(* Logix 5000 project; controller FV vendor 1 type 14 code 217 rev 31.11; software revision 31.00; part 18 of 63 *)
(* tags used below, declared in another part *)
   CheckTimeMask : INT;
   CWD : CHECKWORD_FLAGS;
   Delphi_Does_Eng_Func : BOOL;
   FR_AUDI1 : PlantItem;   // AUDI1
   FR_B240 : INT[255];   // DEBOUNCE Debounce Flags
   FR_BEACON1 : PlantItem;   // BEACON1
   FR_FV26_VA01 : PlantItem;   // FV26_VA01
   FR_FV27_VA01 : PlantItem;   // FV27_VA01
   FR_FV28_V : PlantItem;   // FV28_V
   FR_FV28_VA01 : PlantItem;   // FV28_VA01
   FR_FVS_P01 : PlantItem;   // FVS_P01
   FR_N14 : INT[265];   // MVFV CIP Comms to MVFV CIP Un it PLC
   FR_N140 : INT[265];   // CIP
   FR_N255 : INT[265];   // CHECKWORDS
   FR_N26 : INT[265];   // FV26
   FR_N27 : INT[265];   // FV27
   FR_N28 : INT[265];   // FV28
   FR_N29 : INT[265];   // FV29
   FR_N30 : INT[265];   // FV30
   FR_N31 : INT[265];   // FV31
   FR_N99 : INT[265];   // COMMENT Comment Lines
   FR_R3_SW3_1 : PlantItem;   // R3_SW3_1
   FR_R3_SW3_2 : PlantItem;   // R3_SW3_2
   FR_R3_SW3_3 : PlantItem;   // R3_SW3_3
   FR_T144 : TIMER[255];   // CIP
   FR_VB4_AV20 : PlantItem;   // VB4_AV20
   FR_VB4_AV22 : PlantItem;   // VB4_AV22
   FR_YP1_CIP : PlantItem;   // YP1_CIP
   FR_YP2_CIP : PlantItem;   // YP2_CIP
   FR_YP3_CIP : PlantItem;   // YP3_CIP
   TempChecktime : DINT;
(* FR_Common, continued *)

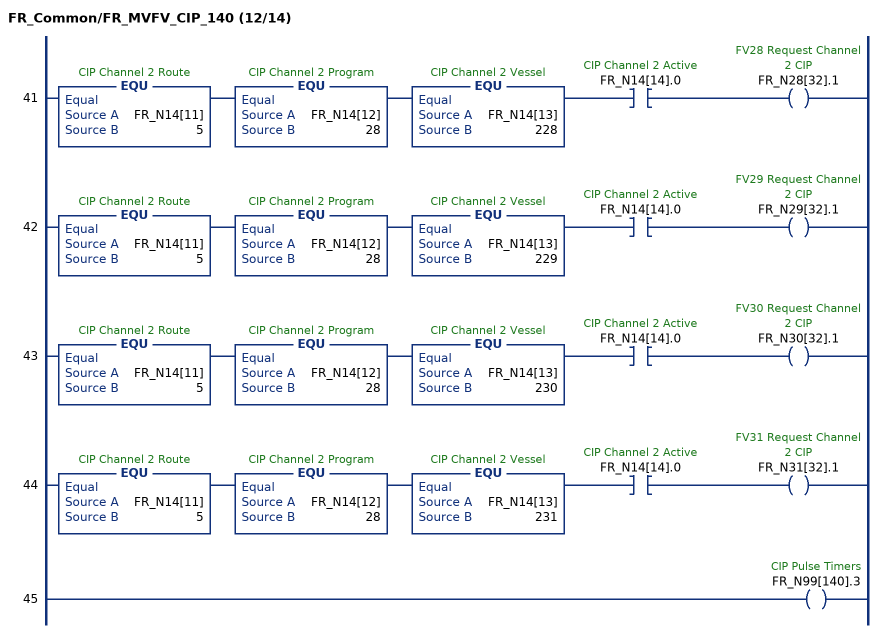
   [picture p297: FR_Common/FR_MVFV_CIP_140 rungs 41-45]
   41: EQU(FR_N14[11],5)EQU(FR_N14[12],28)EQU(FR_N14[13],228)XIC(FR_N14[14].0)OTE(FR_N28[32].1);
   42: EQU(FR_N14[11],5)EQU(FR_N14[12],28)EQU(FR_N14[13],229)XIC(FR_N14[14].0)OTE(FR_N29[32].1);
   43: EQU(FR_N14[11],5)EQU(FR_N14[12],28)EQU(FR_N14[13],230)XIC(FR_N14[14].0)OTE(FR_N30[32].1);
   44: EQU(FR_N14[11],5)EQU(FR_N14[12],28)EQU(FR_N14[13],231)XIC(FR_N14[14].0)OTE(FR_N31[32].1);
   45: OTE(FR_N99[140].3);
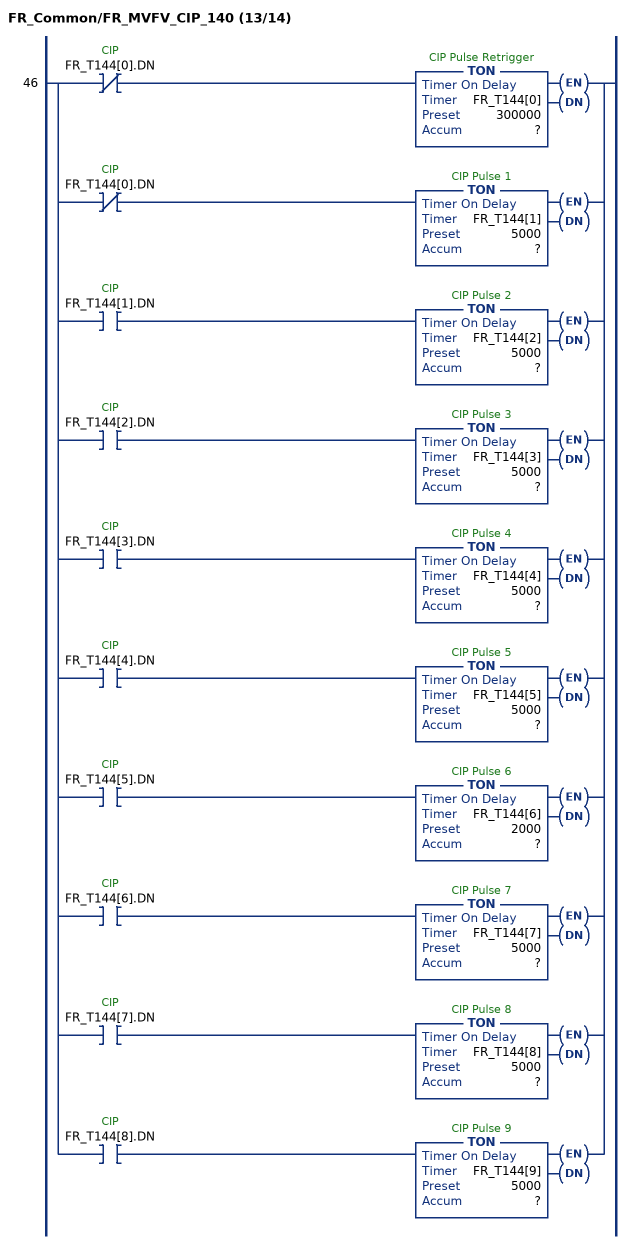
   46: [XIO(FR_T144[0].DN) TON(FR_T144[0],?,?) ,XIO(FR_T144[0].DN) TON(FR_T144[1],?,?) ,XIC(FR_T144[1].DN) TON(FR_T144[2],?,?) ,XIC(FR_T144[2].DN) TON(FR_T144[3],?,?) ,XIC(FR_T144[3].DN) TON(FR_T144[4],?,?) ,XIC(FR_T144[4].DN) TON(FR_T144[5],?,?) ,XIC(FR_T144[5].DN) TON(FR_T144[6],?,?) ,XIC(FR_T144[6].DN) TON(FR_T144[7],?,?) ,XIC(FR_T144[7].DN) TON(FR_T144[8],?,?) ,XIC(FR_T144[8].DN) TON(FR_T144[9],?,?) ];
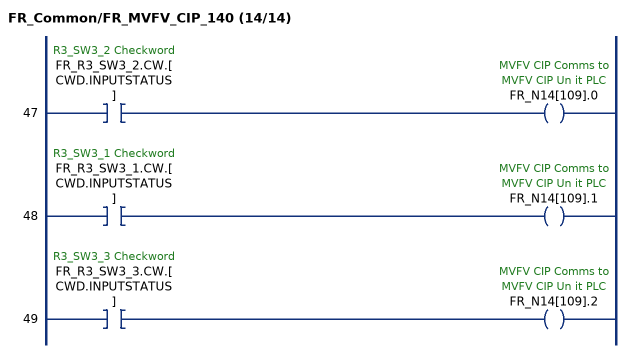
   47: XIC(FR_R3_SW3_2.CW.[CWD.INPUTSTATUS])OTE(FR_N14[109].0);
   48: XIC(FR_R3_SW3_1.CW.[CWD.INPUTSTATUS])OTE(FR_N14[109].1);
   49: XIC(FR_R3_SW3_3.CW.[CWD.INPUTSTATUS])OTE(FR_N14[109].2);
END_ROUTINE

ROUTINE FR_MVFV_CIP_O_141   (* ladder *)
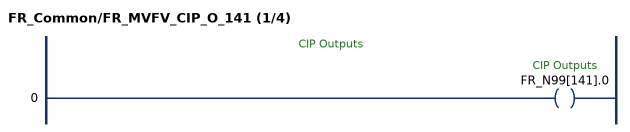
   // CIP Outputs
   0: OTE(FR_N99[141].0);
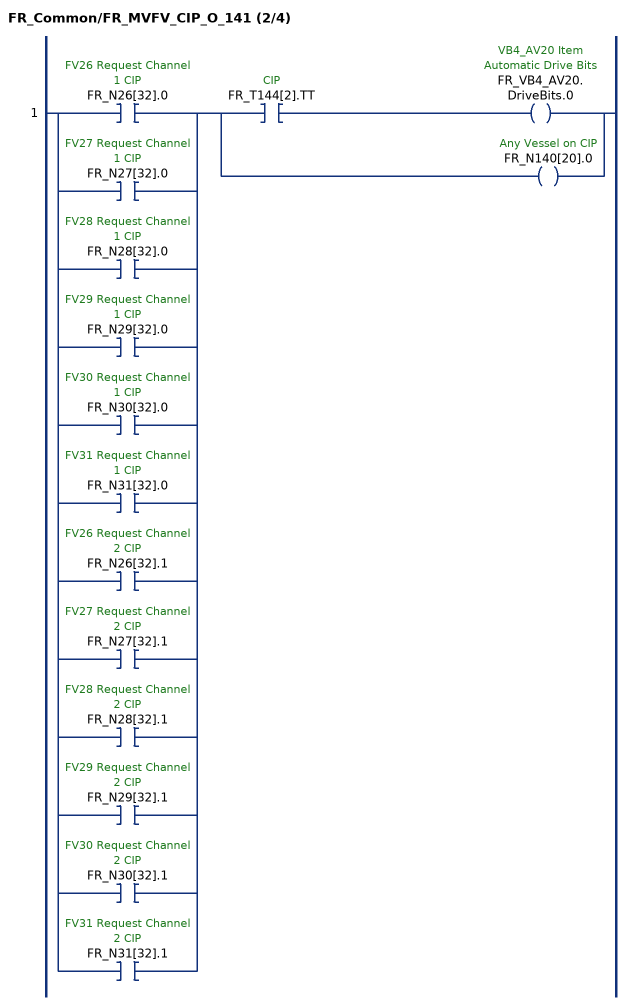
   1: [XIC(FR_N26[32].0) ,XIC(FR_N27[32].0) ,XIC(FR_N28[32].0) ,XIC(FR_N29[32].0) ,XIC(FR_N30[32].0) ,XIC(FR_N31[32].0) ,XIC(FR_N26[32].1) ,XIC(FR_N27[32].1) ,XIC(FR_N28[32].1) ,XIC(FR_N29[32].1) ,XIC(FR_N30[32].1) ,XIC(FR_N31[32].1) ][XIC(FR_T144[2].TT) OTE(FR_VB4_AV20.DriveBits.0) ,OTE(FR_N140[20].0) ];
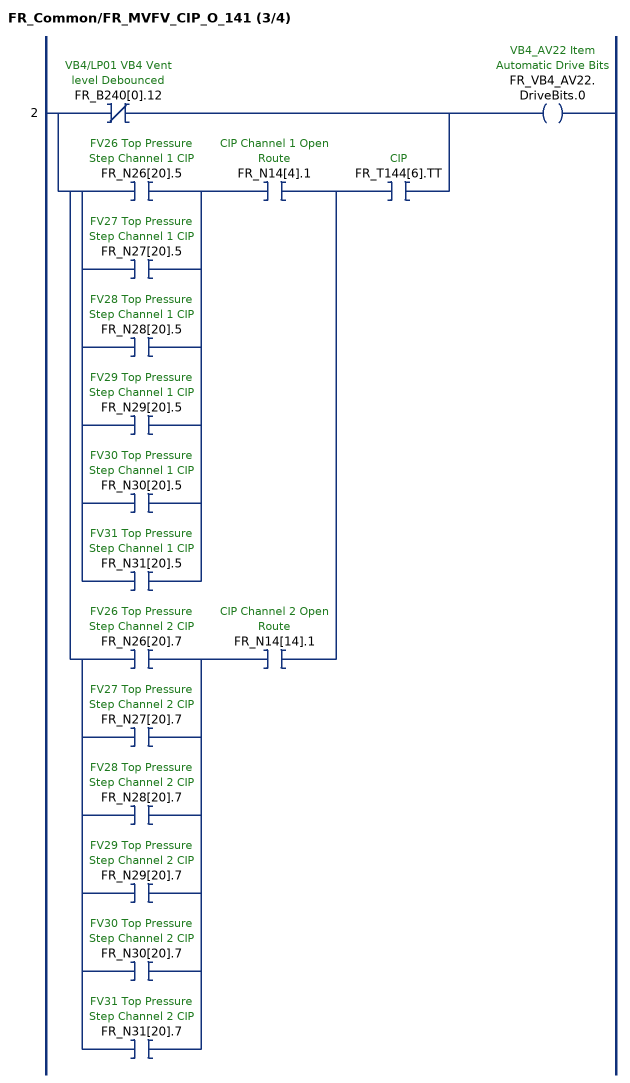
   2: [XIO(FR_B240[0].12) ,[[XIC(FR_N26[20].5) ,XIC(FR_N27[20].5) ,XIC(FR_N28[20].5) ,XIC(FR_N29[20].5) ,XIC(FR_N30[20].5) ,XIC(FR_N31[20].5) ] XIC(FR_N14[4].1) ,[XIC(FR_N26[20].7) ,XIC(FR_N27[20].7) ,XIC(FR_N28[20].7) ,XIC(FR_N29[20].7) ,XIC(FR_N30[20].7) ,XIC(FR_N31[20].7) ] XIC(FR_N14[14].1) ] XIC(FR_T144[6].TT) ]OTE(FR_VB4_AV22.DriveBits.0);
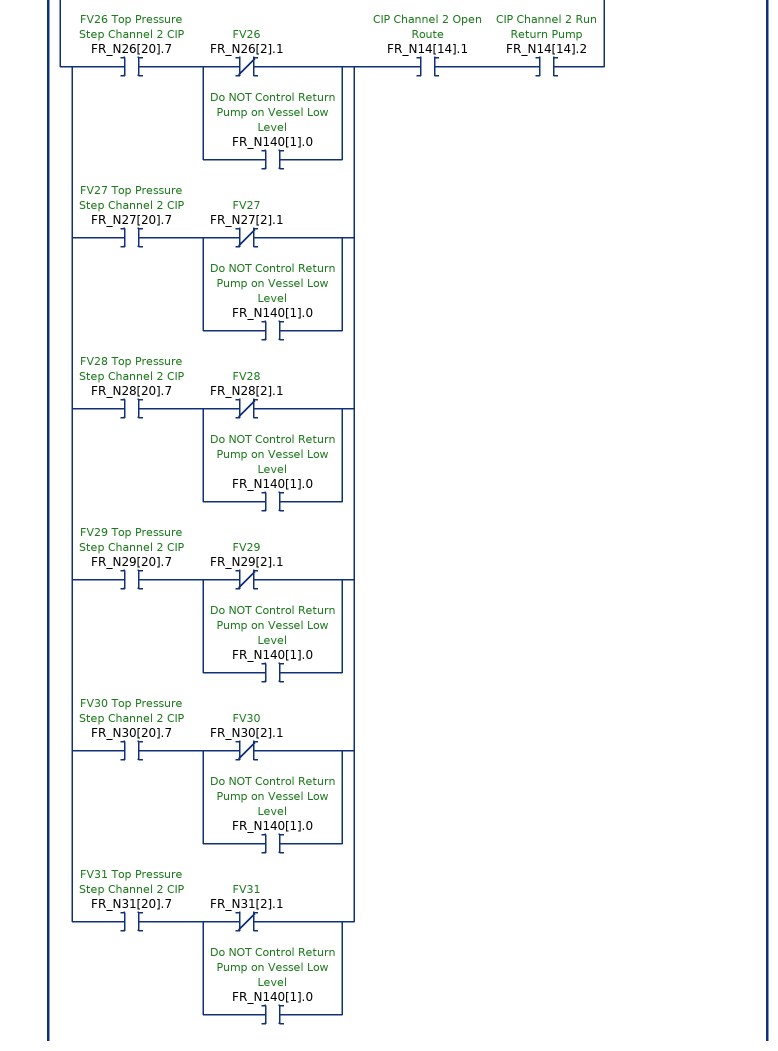
   3: [[XIC(FR_N26[20].5) [XIO(FR_N26[2].1) ,XIC(FR_N140[1].0) ] ,XIC(FR_N27[20].5) [XIO(FR_N27[2].1) ,XIC(FR_N140[1].0) ] ,XIC(FR_N28[20].5) [XIO(FR_N28[2].1) ,XIC(FR_N140[1].0) ] ,XIC(FR_N29[20].5) [XIO(FR_N29[2].1) ,XIC(FR_N140[1].0) ] ,XIC(FR_N30[20].5) [XIO(FR_N30[2].1) ,XIC(FR_N140[1].0) ] ,XIC(FR_N31[20].5) [XIO(FR_N31[2].1) ,XIC(FR_N140[1].0) ] ] XIC(FR_N14[4].1) XIC(FR_N14[4].2) ,[XIC(FR_N26[20].7) [XIO(FR_N26[2].1) ,XIC(FR_N140[1].0) ] ,XIC(FR_N27[20].7) [XIO(FR_N27[2].1) ,XIC(FR_N140[1].0) ] ,XIC(FR_N28[20].7) [XIO(FR_N28[2].1) ,XIC(FR_N140[1].0) ] ,XIC(FR_N29[20].7) [XIO(FR_N29[2].1) ,XIC(FR_N140[1].0) ] ,XIC(FR_N30[20].7) [XIO(FR_N30[2].1) ,XIC(FR_N140[1].0) ] ,XIC(FR_N31[20].7) [XIO(FR_N31[2].1) ,XIC(FR_N140[1].0) ] ] XIC(FR_N14[14].1) XIC(FR_N14[14].2) ]OTE(FR_FVS_P01.DriveBits.0);
END_ROUTINE

ROUTINE FR_Old_Checkword_Relaying   (* ladder *)
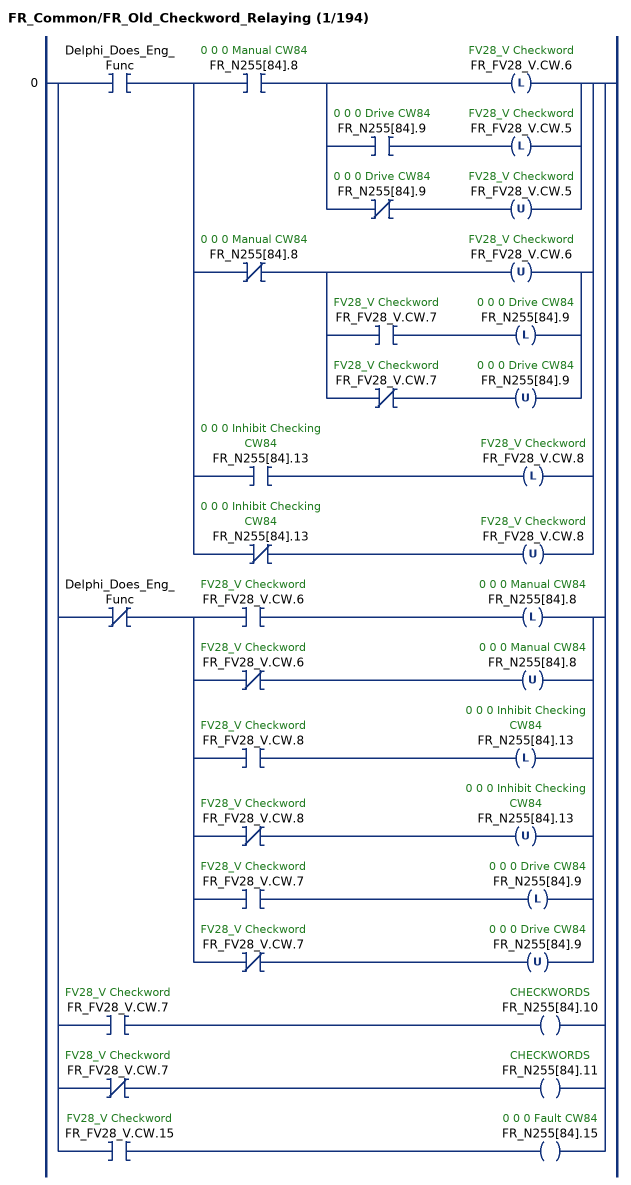
   0: [XIC(Delphi_Does_Eng_Func) [[XIC(FR_N255[84].8) [OTL(FR_FV28_V.CW.6) ,XIC(FR_N255[84].9) OTL(FR_FV28_V.CW.5) ,XIO(FR_N255[84].9) OTU(FR_FV28_V.CW.5) ] ,XIO(FR_N255[84].8) [OTU(FR_FV28_V.CW.6) ,[XIC(FR_FV28_V.CW.7) OTL(FR_N255[84].9) ,XIO(FR_FV28_V.CW.7) OTU(FR_N255[84].9) ] ] ] ,[XIC(FR_N255[84].13) OTL(FR_FV28_V.CW.8) ,XIO(FR_N255[84].13) OTU(FR_FV28_V.CW.8) ] ] ,XIO(Delphi_Does_Eng_Func) [[XIC(FR_FV28_V.CW.6) OTL(FR_N255[84].8) ,XIO(FR_FV28_V.CW.6) OTU(FR_N255[84].8) ] ,[XIC(FR_FV28_V.CW.8) OTL(FR_N255[84].13) ,XIO(FR_FV28_V.CW.8) OTU(FR_N255[84].13) ] ,[XIC(FR_FV28_V.CW.7) OTL(FR_N255[84].9) ,XIO(FR_FV28_V.CW.7) OTU(FR_N255[84].9) ] ] ,XIC(FR_FV28_V.CW.7) OTE(FR_N255[84].10) ,XIO(FR_FV28_V.CW.7) OTE(FR_N255[84].11) ,XIC(FR_FV28_V.CW.15) OTE(FR_N255[84].15) ];
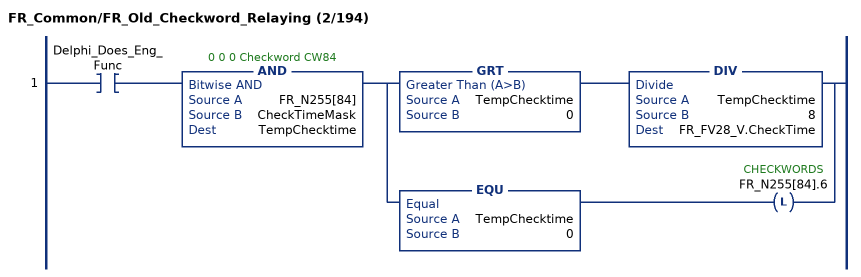
   1: XIC(Delphi_Does_Eng_Func)AND(FR_N255[84],CheckTimeMask,TempChecktime)[GRT(TempChecktime,0) DIV(TempChecktime,8,FR_FV28_V.CheckTime) ,EQU(TempChecktime,0) OTL(FR_N255[84].6) ];
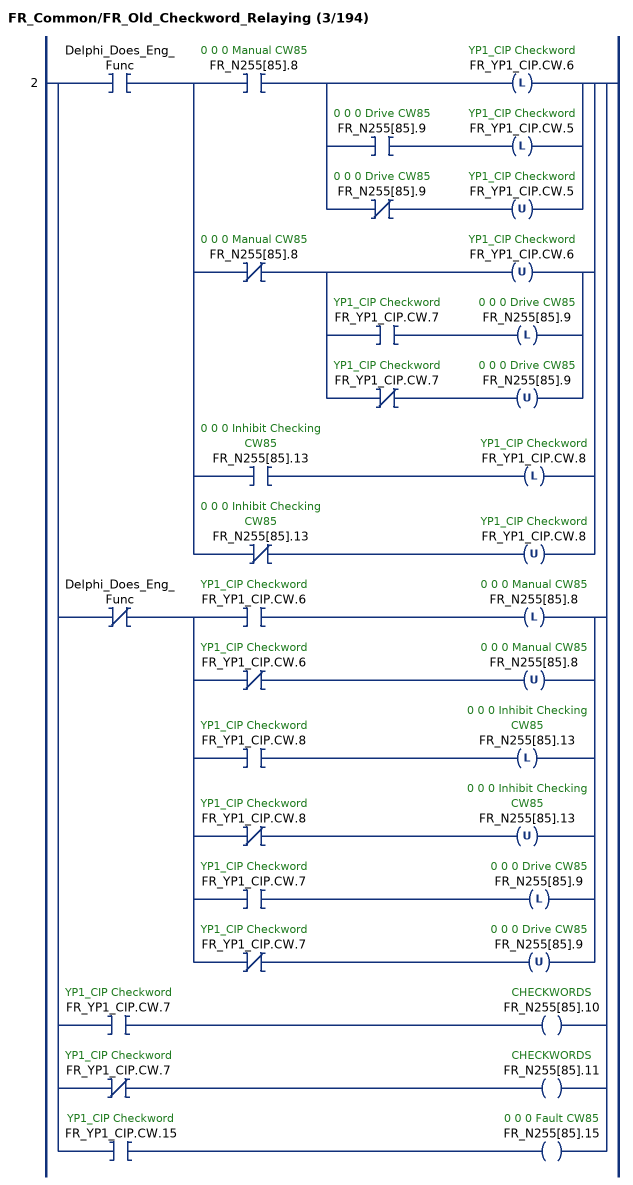
   2: [XIC(Delphi_Does_Eng_Func) [[XIC(FR_N255[85].8) [OTL(FR_YP1_CIP.CW.6) ,XIC(FR_N255[85].9) OTL(FR_YP1_CIP.CW.5) ,XIO(FR_N255[85].9) OTU(FR_YP1_CIP.CW.5) ] ,XIO(FR_N255[85].8) [OTU(FR_YP1_CIP.CW.6) ,[XIC(FR_YP1_CIP.CW.7) OTL(FR_N255[85].9) ,XIO(FR_YP1_CIP.CW.7) OTU(FR_N255[85].9) ] ] ] ,[XIC(FR_N255[85].13) OTL(FR_YP1_CIP.CW.8) ,XIO(FR_N255[85].13) OTU(FR_YP1_CIP.CW.8) ] ] ,XIO(Delphi_Does_Eng_Func) [[XIC(FR_YP1_CIP.CW.6) OTL(FR_N255[85].8) ,XIO(FR_YP1_CIP.CW.6) OTU(FR_N255[85].8) ] ,[XIC(FR_YP1_CIP.CW.8) OTL(FR_N255[85].13) ,XIO(FR_YP1_CIP.CW.8) OTU(FR_N255[85].13) ] ,[XIC(FR_YP1_CIP.CW.7) OTL(FR_N255[85].9) ,XIO(FR_YP1_CIP.CW.7) OTU(FR_N255[85].9) ] ] ,XIC(FR_YP1_CIP.CW.7) OTE(FR_N255[85].10) ,XIO(FR_YP1_CIP.CW.7) OTE(FR_N255[85].11) ,XIC(FR_YP1_CIP.CW.15) OTE(FR_N255[85].15) ];
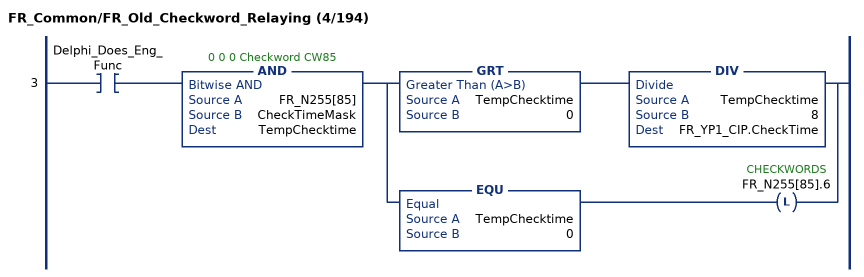
   3: XIC(Delphi_Does_Eng_Func)AND(FR_N255[85],CheckTimeMask,TempChecktime)[GRT(TempChecktime,0) DIV(TempChecktime,8,FR_YP1_CIP.CheckTime) ,EQU(TempChecktime,0) OTL(FR_N255[85].6) ];
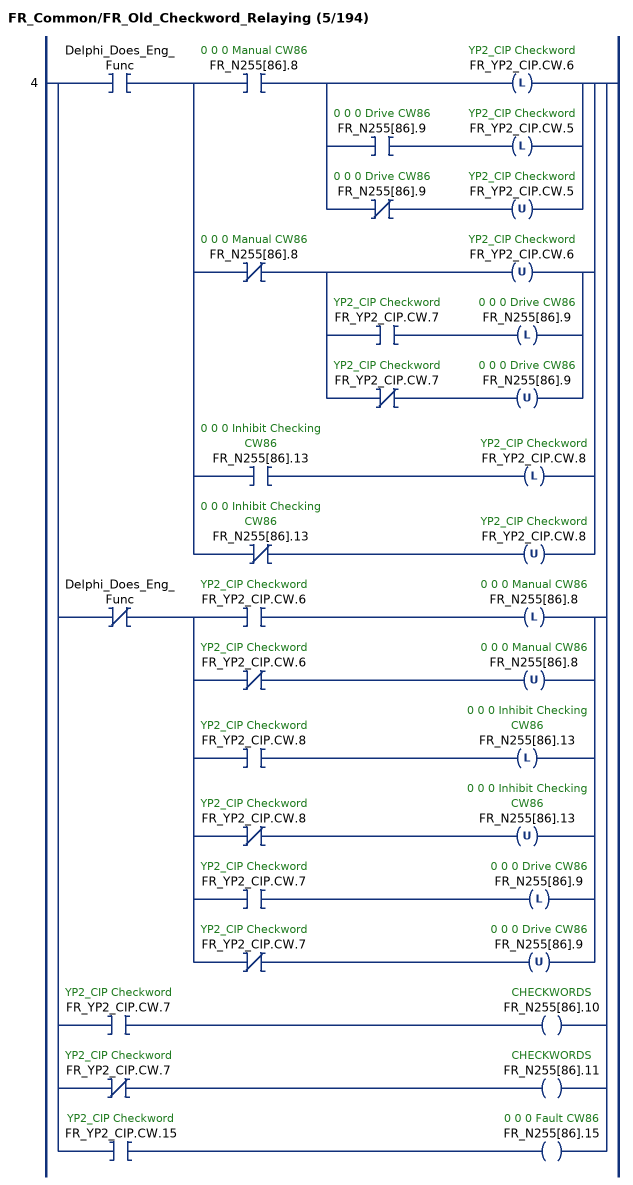
   4: [XIC(Delphi_Does_Eng_Func) [[XIC(FR_N255[86].8) [OTL(FR_YP2_CIP.CW.6) ,XIC(FR_N255[86].9) OTL(FR_YP2_CIP.CW.5) ,XIO(FR_N255[86].9) OTU(FR_YP2_CIP.CW.5) ] ,XIO(FR_N255[86].8) [OTU(FR_YP2_CIP.CW.6) ,[XIC(FR_YP2_CIP.CW.7) OTL(FR_N255[86].9) ,XIO(FR_YP2_CIP.CW.7) OTU(FR_N255[86].9) ] ] ] ,[XIC(FR_N255[86].13) OTL(FR_YP2_CIP.CW.8) ,XIO(FR_N255[86].13) OTU(FR_YP2_CIP.CW.8) ] ] ,XIO(Delphi_Does_Eng_Func) [[XIC(FR_YP2_CIP.CW.6) OTL(FR_N255[86].8) ,XIO(FR_YP2_CIP.CW.6) OTU(FR_N255[86].8) ] ,[XIC(FR_YP2_CIP.CW.8) OTL(FR_N255[86].13) ,XIO(FR_YP2_CIP.CW.8) OTU(FR_N255[86].13) ] ,[XIC(FR_YP2_CIP.CW.7) OTL(FR_N255[86].9) ,XIO(FR_YP2_CIP.CW.7) OTU(FR_N255[86].9) ] ] ,XIC(FR_YP2_CIP.CW.7) OTE(FR_N255[86].10) ,XIO(FR_YP2_CIP.CW.7) OTE(FR_N255[86].11) ,XIC(FR_YP2_CIP.CW.15) OTE(FR_N255[86].15) ];
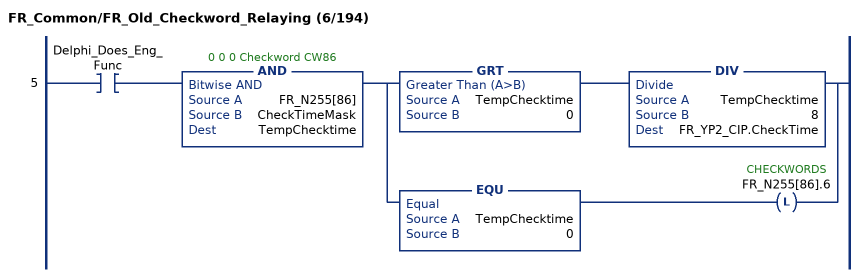
   5: XIC(Delphi_Does_Eng_Func)AND(FR_N255[86],CheckTimeMask,TempChecktime)[GRT(TempChecktime,0) DIV(TempChecktime,8,FR_YP2_CIP.CheckTime) ,EQU(TempChecktime,0) OTL(FR_N255[86].6) ];
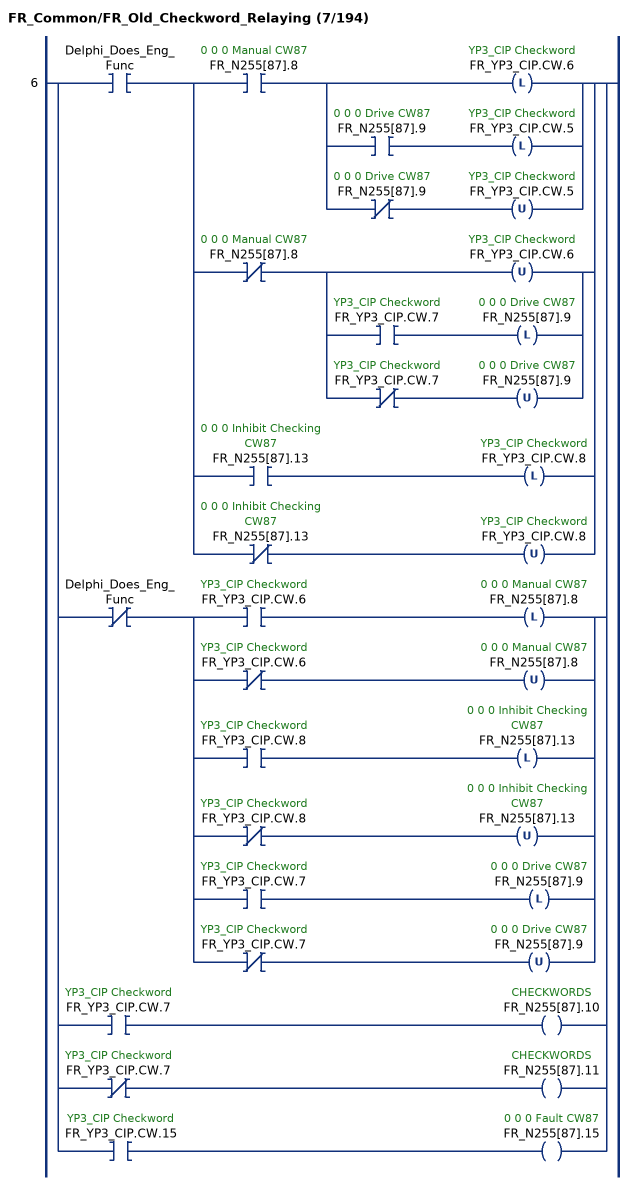
   6: [XIC(Delphi_Does_Eng_Func) [[XIC(FR_N255[87].8) [OTL(FR_YP3_CIP.CW.6) ,XIC(FR_N255[87].9) OTL(FR_YP3_CIP.CW.5) ,XIO(FR_N255[87].9) OTU(FR_YP3_CIP.CW.5) ] ,XIO(FR_N255[87].8) [OTU(FR_YP3_CIP.CW.6) ,[XIC(FR_YP3_CIP.CW.7) OTL(FR_N255[87].9) ,XIO(FR_YP3_CIP.CW.7) OTU(FR_N255[87].9) ] ] ] ,[XIC(FR_N255[87].13) OTL(FR_YP3_CIP.CW.8) ,XIO(FR_N255[87].13) OTU(FR_YP3_CIP.CW.8) ] ] ,XIO(Delphi_Does_Eng_Func) [[XIC(FR_YP3_CIP.CW.6) OTL(FR_N255[87].8) ,XIO(FR_YP3_CIP.CW.6) OTU(FR_N255[87].8) ] ,[XIC(FR_YP3_CIP.CW.8) OTL(FR_N255[87].13) ,XIO(FR_YP3_CIP.CW.8) OTU(FR_N255[87].13) ] ,[XIC(FR_YP3_CIP.CW.7) OTL(FR_N255[87].9) ,XIO(FR_YP3_CIP.CW.7) OTU(FR_N255[87].9) ] ] ,XIC(FR_YP3_CIP.CW.7) OTE(FR_N255[87].10) ,XIO(FR_YP3_CIP.CW.7) OTE(FR_N255[87].11) ,XIC(FR_YP3_CIP.CW.15) OTE(FR_N255[87].15) ];
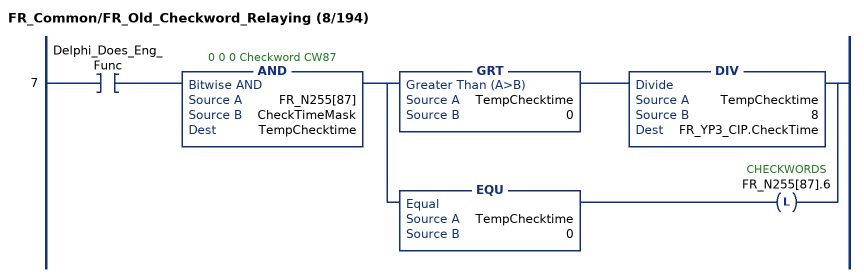
   7: XIC(Delphi_Does_Eng_Func)AND(FR_N255[87],CheckTimeMask,TempChecktime)[GRT(TempChecktime,0) DIV(TempChecktime,8,FR_YP3_CIP.CheckTime) ,EQU(TempChecktime,0) OTL(FR_N255[87].6) ];
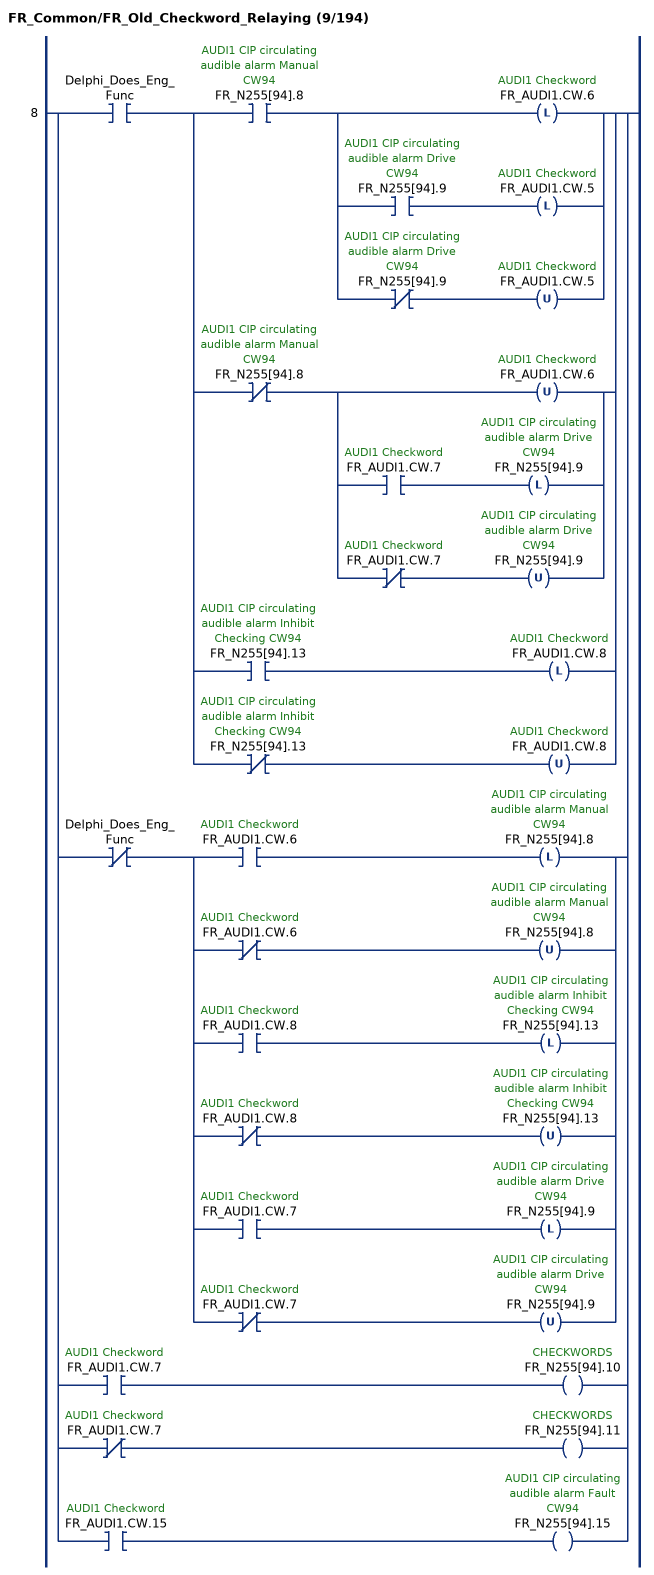
   8: [XIC(Delphi_Does_Eng_Func) [[XIC(FR_N255[94].8) [OTL(FR_AUDI1.CW.6) ,XIC(FR_N255[94].9) OTL(FR_AUDI1.CW.5) ,XIO(FR_N255[94].9) OTU(FR_AUDI1.CW.5) ] ,XIO(FR_N255[94].8) [OTU(FR_AUDI1.CW.6) ,[XIC(FR_AUDI1.CW.7) OTL(FR_N255[94].9) ,XIO(FR_AUDI1.CW.7) OTU(FR_N255[94].9) ] ] ] ,[XIC(FR_N255[94].13) OTL(FR_AUDI1.CW.8) ,XIO(FR_N255[94].13) OTU(FR_AUDI1.CW.8) ] ] ,XIO(Delphi_Does_Eng_Func) [[XIC(FR_AUDI1.CW.6) OTL(FR_N255[94].8) ,XIO(FR_AUDI1.CW.6) OTU(FR_N255[94].8) ] ,[XIC(FR_AUDI1.CW.8) OTL(FR_N255[94].13) ,XIO(FR_AUDI1.CW.8) OTU(FR_N255[94].13) ] ,[XIC(FR_AUDI1.CW.7) OTL(FR_N255[94].9) ,XIO(FR_AUDI1.CW.7) OTU(FR_N255[94].9) ] ] ,XIC(FR_AUDI1.CW.7) OTE(FR_N255[94].10) ,XIO(FR_AUDI1.CW.7) OTE(FR_N255[94].11) ,XIC(FR_AUDI1.CW.15) OTE(FR_N255[94].15) ];
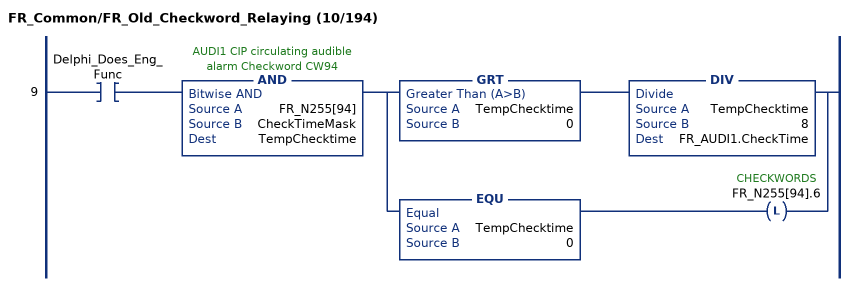
   9: XIC(Delphi_Does_Eng_Func)AND(FR_N255[94],CheckTimeMask,TempChecktime)[GRT(TempChecktime,0) DIV(TempChecktime,8,FR_AUDI1.CheckTime) ,EQU(TempChecktime,0) OTL(FR_N255[94].6) ];
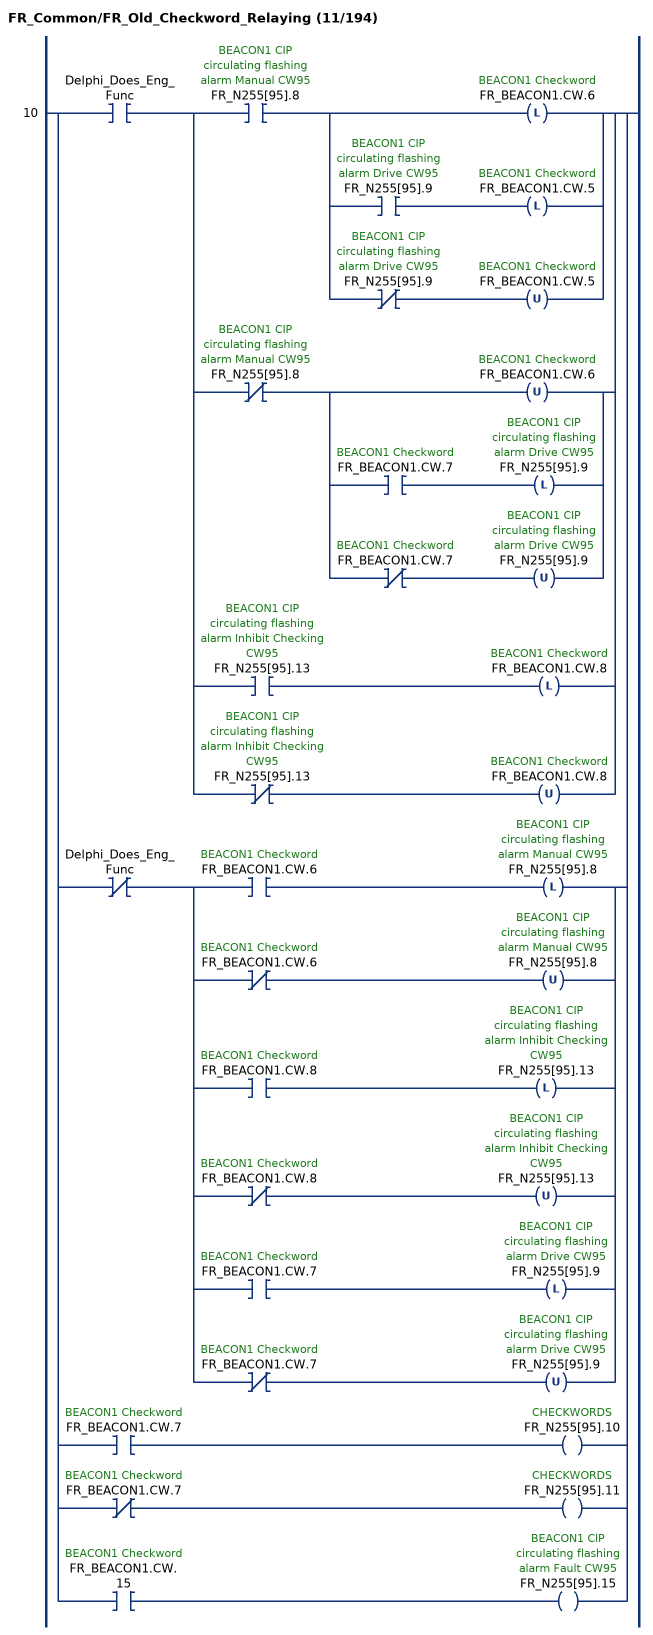
   10: [XIC(Delphi_Does_Eng_Func) [[XIC(FR_N255[95].8) [OTL(FR_BEACON1.CW.6) ,XIC(FR_N255[95].9) OTL(FR_BEACON1.CW.5) ,XIO(FR_N255[95].9) OTU(FR_BEACON1.CW.5) ] ,XIO(FR_N255[95].8) [OTU(FR_BEACON1.CW.6) ,[XIC(FR_BEACON1.CW.7) OTL(FR_N255[95].9) ,XIO(FR_BEACON1.CW.7) OTU(FR_N255[95].9) ] ] ] ,[XIC(FR_N255[95].13) OTL(FR_BEACON1.CW.8) ,XIO(FR_N255[95].13) OTU(FR_BEACON1.CW.8) ] ] ,XIO(Delphi_Does_Eng_Func) [[XIC(FR_BEACON1.CW.6) OTL(FR_N255[95].8) ,XIO(FR_BEACON1.CW.6) OTU(FR_N255[95].8) ] ,[XIC(FR_BEACON1.CW.8) OTL(FR_N255[95].13) ,XIO(FR_BEACON1.CW.8) OTU(FR_N255[95].13) ] ,[XIC(FR_BEACON1.CW.7) OTL(FR_N255[95].9) ,XIO(FR_BEACON1.CW.7) OTU(FR_N255[95].9) ] ] ,XIC(FR_BEACON1.CW.7) OTE(FR_N255[95].10) ,XIO(FR_BEACON1.CW.7) OTE(FR_N255[95].11) ,XIC(FR_BEACON1.CW.15) OTE(FR_N255[95].15) ];
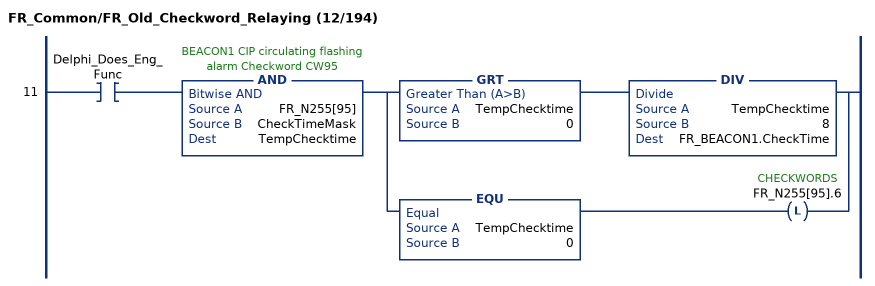
   11: XIC(Delphi_Does_Eng_Func)AND(FR_N255[95],CheckTimeMask,TempChecktime)[GRT(TempChecktime,0) DIV(TempChecktime,8,FR_BEACON1.CheckTime) ,EQU(TempChecktime,0) OTL(FR_N255[95].6) ];
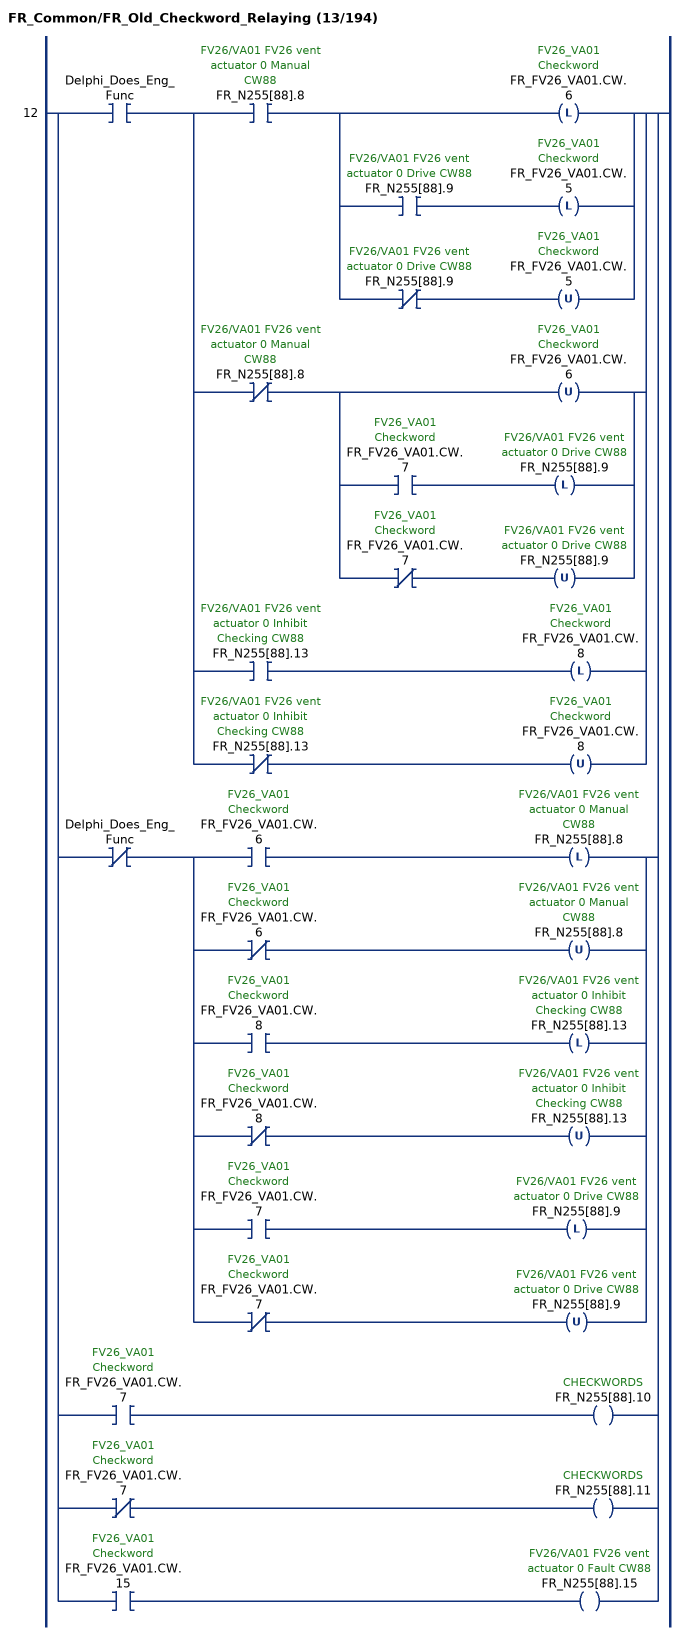
   12: [XIC(Delphi_Does_Eng_Func) [[XIC(FR_N255[88].8) [OTL(FR_FV26_VA01.CW.6) ,XIC(FR_N255[88].9) OTL(FR_FV26_VA01.CW.5) ,XIO(FR_N255[88].9) OTU(FR_FV26_VA01.CW.5) ] ,XIO(FR_N255[88].8) [OTU(FR_FV26_VA01.CW.6) ,[XIC(FR_FV26_VA01.CW.7) OTL(FR_N255[88].9) ,XIO(FR_FV26_VA01.CW.7) OTU(FR_N255[88].9) ] ] ] ,[XIC(FR_N255[88].13) OTL(FR_FV26_VA01.CW.8) ,XIO(FR_N255[88].13) OTU(FR_FV26_VA01.CW.8) ] ] ,XIO(Delphi_Does_Eng_Func) [[XIC(FR_FV26_VA01.CW.6) OTL(FR_N255[88].8) ,XIO(FR_FV26_VA01.CW.6) OTU(FR_N255[88].8) ] ,[XIC(FR_FV26_VA01.CW.8) OTL(FR_N255[88].13) ,XIO(FR_FV26_VA01.CW.8) OTU(FR_N255[88].13) ] ,[XIC(FR_FV26_VA01.CW.7) OTL(FR_N255[88].9) ,XIO(FR_FV26_VA01.CW.7) OTU(FR_N255[88].9) ] ] ,XIC(FR_FV26_VA01.CW.7) OTE(FR_N255[88].10) ,XIO(FR_FV26_VA01.CW.7) OTE(FR_N255[88].11) ,XIC(FR_FV26_VA01.CW.15) OTE(FR_N255[88].15) ];
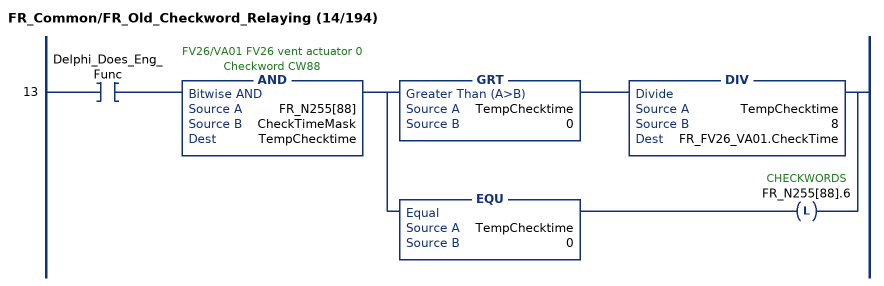
   13: XIC(Delphi_Does_Eng_Func)AND(FR_N255[88],CheckTimeMask,TempChecktime)[GRT(TempChecktime,0) DIV(TempChecktime,8,FR_FV26_VA01.CheckTime) ,EQU(TempChecktime,0) OTL(FR_N255[88].6) ];
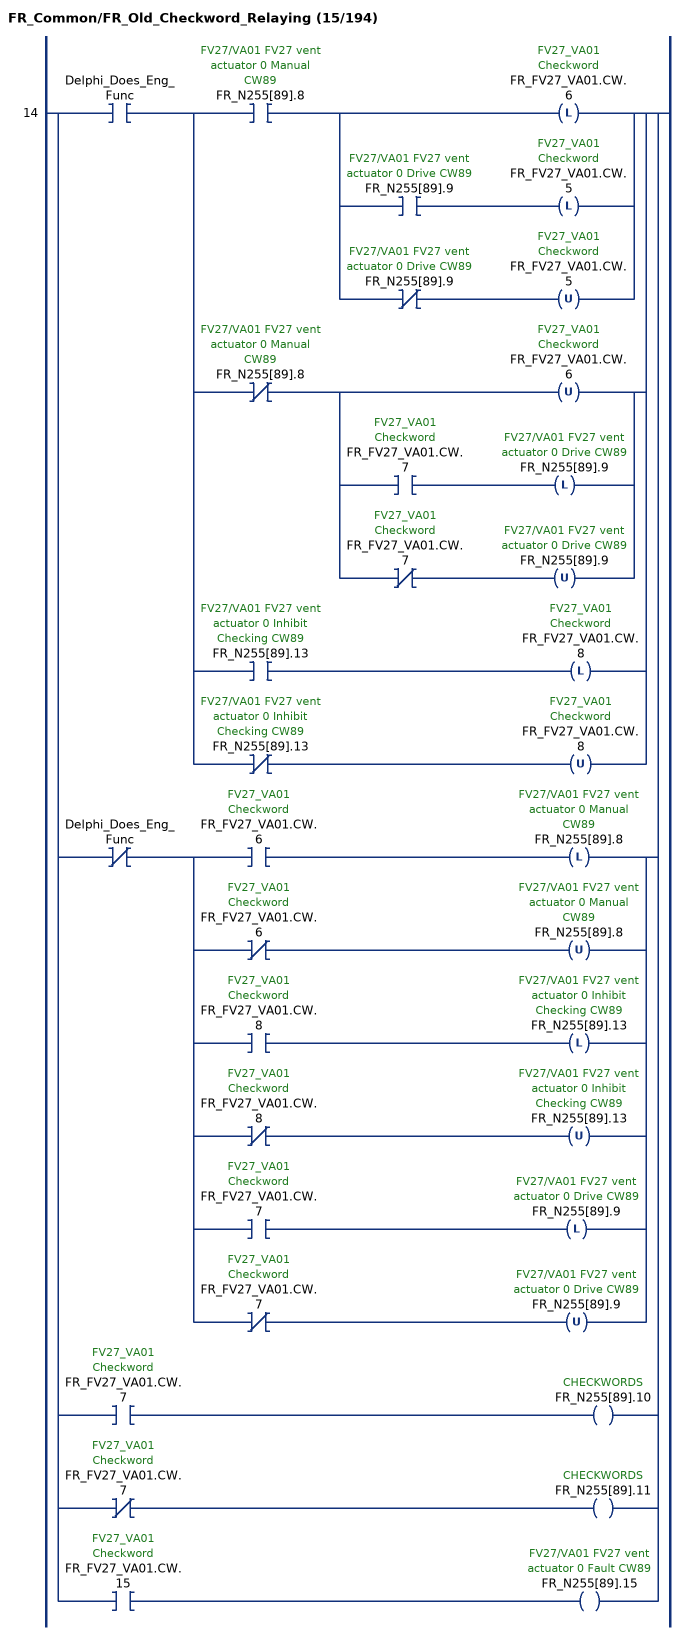
   14: [XIC(Delphi_Does_Eng_Func) [[XIC(FR_N255[89].8) [OTL(FR_FV27_VA01.CW.6) ,XIC(FR_N255[89].9) OTL(FR_FV27_VA01.CW.5) ,XIO(FR_N255[89].9) OTU(FR_FV27_VA01.CW.5) ] ,XIO(FR_N255[89].8) [OTU(FR_FV27_VA01.CW.6) ,[XIC(FR_FV27_VA01.CW.7) OTL(FR_N255[89].9) ,XIO(FR_FV27_VA01.CW.7) OTU(FR_N255[89].9) ] ] ] ,[XIC(FR_N255[89].13) OTL(FR_FV27_VA01.CW.8) ,XIO(FR_N255[89].13) OTU(FR_FV27_VA01.CW.8) ] ] ,XIO(Delphi_Does_Eng_Func) [[XIC(FR_FV27_VA01.CW.6) OTL(FR_N255[89].8) ,XIO(FR_FV27_VA01.CW.6) OTU(FR_N255[89].8) ] ,[XIC(FR_FV27_VA01.CW.8) OTL(FR_N255[89].13) ,XIO(FR_FV27_VA01.CW.8) OTU(FR_N255[89].13) ] ,[XIC(FR_FV27_VA01.CW.7) OTL(FR_N255[89].9) ,XIO(FR_FV27_VA01.CW.7) OTU(FR_N255[89].9) ] ] ,XIC(FR_FV27_VA01.CW.7) OTE(FR_N255[89].10) ,XIO(FR_FV27_VA01.CW.7) OTE(FR_N255[89].11) ,XIC(FR_FV27_VA01.CW.15) OTE(FR_N255[89].15) ];
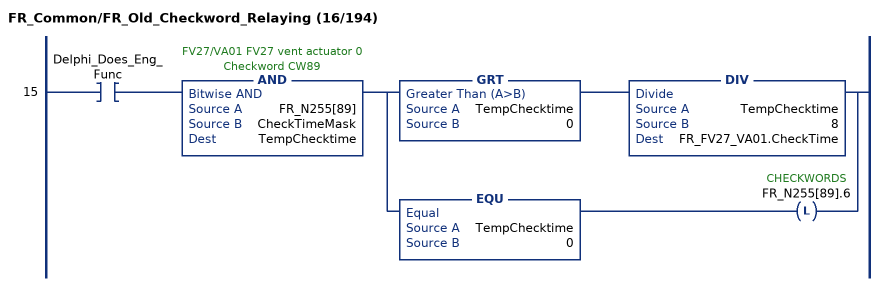
   15: XIC(Delphi_Does_Eng_Func)AND(FR_N255[89],CheckTimeMask,TempChecktime)[GRT(TempChecktime,0) DIV(TempChecktime,8,FR_FV27_VA01.CheckTime) ,EQU(TempChecktime,0) OTL(FR_N255[89].6) ];
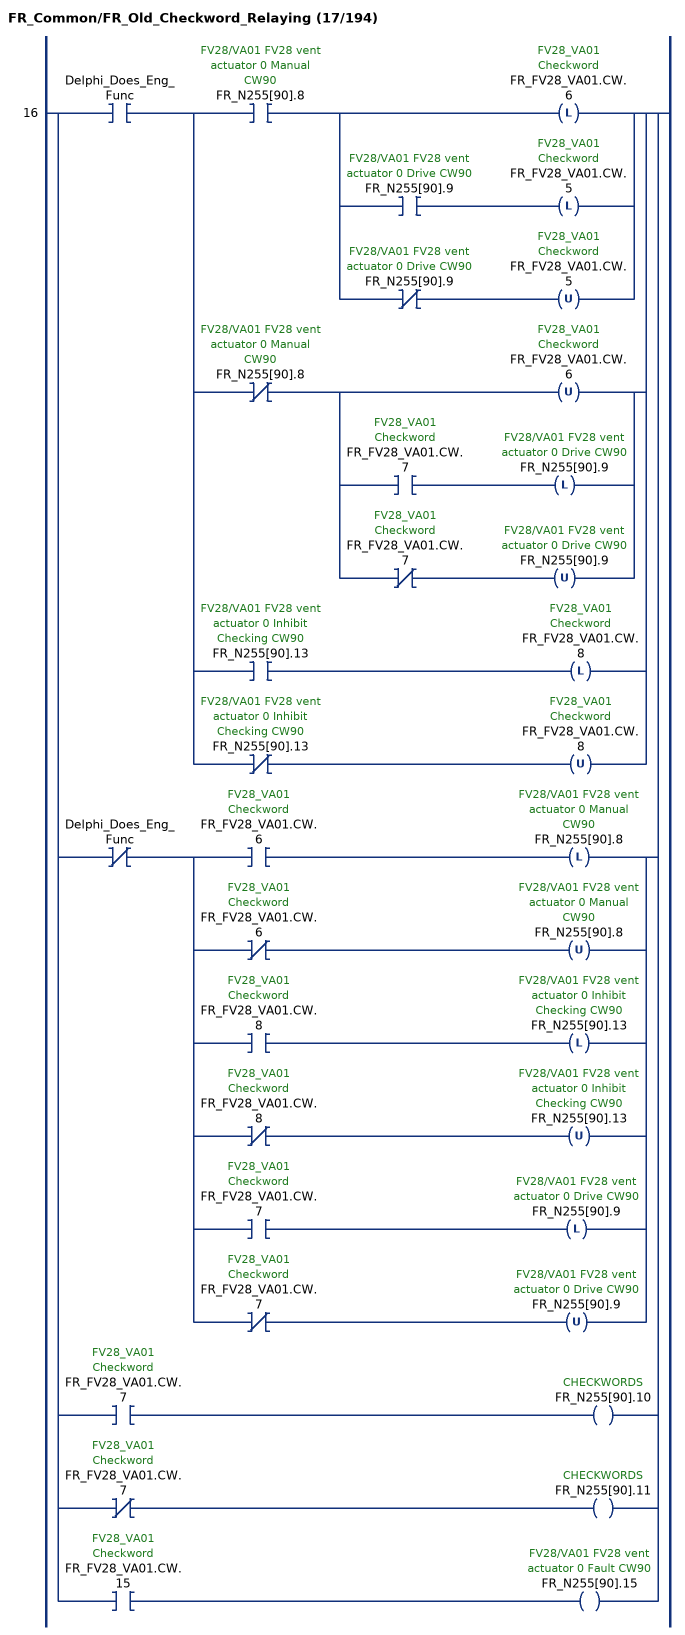
   16: [XIC(Delphi_Does_Eng_Func) [[XIC(FR_N255[90].8) [OTL(FR_FV28_VA01.CW.6) ,XIC(FR_N255[90].9) OTL(FR_FV28_VA01.CW.5) ,XIO(FR_N255[90].9) OTU(FR_FV28_VA01.CW.5) ] ,XIO(FR_N255[90].8) [OTU(FR_FV28_VA01.CW.6) ,[XIC(FR_FV28_VA01.CW.7) OTL(FR_N255[90].9) ,XIO(FR_FV28_VA01.CW.7) OTU(FR_N255[90].9) ] ] ] ,[XIC(FR_N255[90].13) OTL(FR_FV28_VA01.CW.8) ,XIO(FR_N255[90].13) OTU(FR_FV28_VA01.CW.8) ] ] ,XIO(Delphi_Does_Eng_Func) [[XIC(FR_FV28_VA01.CW.6) OTL(FR_N255[90].8) ,XIO(FR_FV28_VA01.CW.6) OTU(FR_N255[90].8) ] ,[XIC(FR_FV28_VA01.CW.8) OTL(FR_N255[90].13) ,XIO(FR_FV28_VA01.CW.8) OTU(FR_N255[90].13) ] ,[XIC(FR_FV28_VA01.CW.7) OTL(FR_N255[90].9) ,XIO(FR_FV28_VA01.CW.7) OTU(FR_N255[90].9) ] ] ,XIC(FR_FV28_VA01.CW.7) OTE(FR_N255[90].10) ,XIO(FR_FV28_VA01.CW.7) OTE(FR_N255[90].11) ,XIC(FR_FV28_VA01.CW.15) OTE(FR_N255[90].15) ];
